(* Logix 5000 project; controller MV vendor 1 type 14 code 217 rev 31.11; software revision 31.00; part 7 of 53 *)
(* tags used below, declared in another part *)
   active : BOOL;
   Ch1_cmd_scan_count : DINT;
   Ch1_DataDelay : TIMER;
   MC_CH1_DRAIN : PlantItem;   // CH1_DRAIN
   MC_CH1_RR : PlantItem;   // CH1_RR
   MC_data_file_value_to_move : DINT;
   MC_N100 : INT[255];   // C1_PLC Channel 1 PLC data
   MC_N101 : INT[255];   // CH1 PC>PLC Channel 1 PC to PLC
   MC_N102 : INT[255];   // CH1 PROG Channel 1 CIP progra m
   MC_N104 : INT[255];   // CH1 REPORT Channel 1 CIP report file
   MC_N108 : INT[255];   // CH1 VDATA Channel 1 CIP progra m validation data
   MC_N120 : INT[255];   // C2 PLC Channel 2 PLC data
   MC_T105 : TIMER[255];   // CH1 TIMERS Channel 1 timers
   MC_T4 : TIMER[255];   // TIMER
(* MC_Common, continued *)

ROUTINE MC_CH1_CMD_101   (* ladder *)
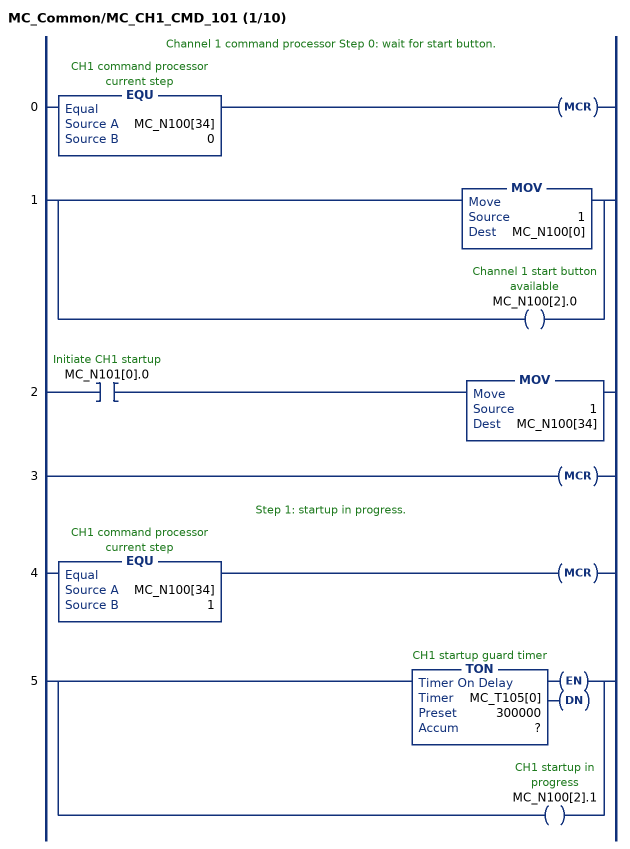
   // Channel 1 command processor Step 0: wait for start button.
   0: EQU(MC_N100[34],0)MCR();
   1: [MOV(1,MC_N100[0]) ,OTE(MC_N100[2].0) ];
   2: XIC(MC_N101[0].0)MOV(1,MC_N100[34]);
   3: MCR();
   // Step 1: startup in progress.
   4: EQU(MC_N100[34],1)MCR();
   5: [TON(MC_T105[0],?,?) ,OTE(MC_N100[2].1) ];
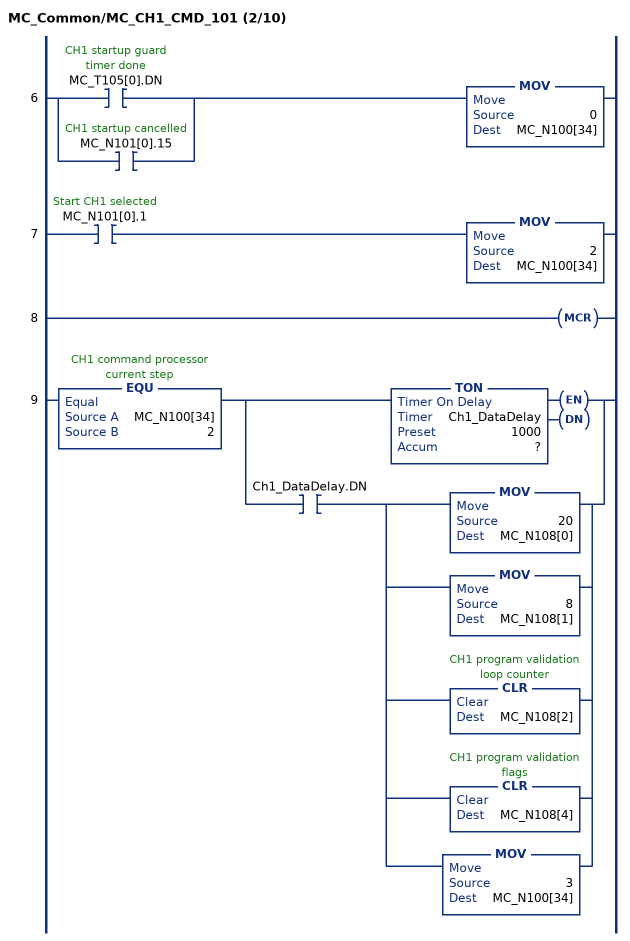
   6: [XIC(MC_T105[0].DN) ,XIC(MC_N101[0].15) ]MOV(0,MC_N100[34]);
   7: XIC(MC_N101[0].1)MOV(2,MC_N100[34]);
   8: MCR();
   9: EQU(MC_N100[34],2)[TON(Ch1_DataDelay,?,?) ,XIC(Ch1_DataDelay.DN) [MOV(20,MC_N108[0]) ,MOV(8,MC_N108[1]) ,CLR(MC_N108[2]) ,CLR(MC_N108[4]) ,MOV(3,MC_N100[34]) ] ];
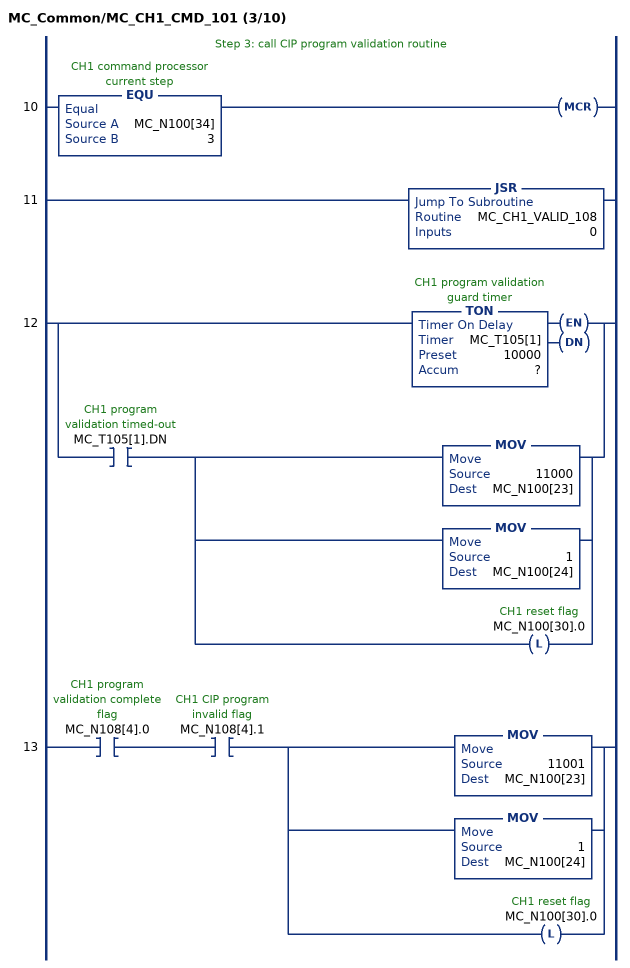
   // Step 3: call CIP program validation routine
   10: EQU(MC_N100[34],3)MCR();
   11: JSR(MC_CH1_VALID_108,0);
   12: [TON(MC_T105[1],?,?) ,XIC(MC_T105[1].DN) [MOV(11000,MC_N100[23]) ,MOV(1,MC_N100[24]) ,OTL(MC_N100[30].0) ] ];
   13: XIC(MC_N108[4].0)XIC(MC_N108[4].1)[MOV(11001,MC_N100[23]) ,MOV(1,MC_N100[24]) ,OTL(MC_N100[30].0) ];
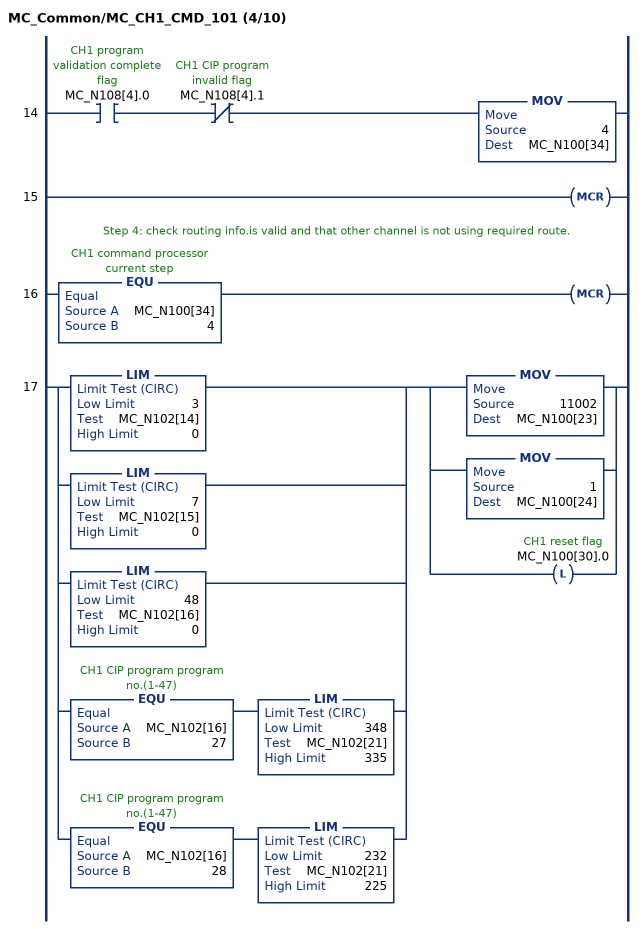
   14: XIC(MC_N108[4].0)XIO(MC_N108[4].1)MOV(4,MC_N100[34]);
   15: MCR();
   // Step 4: check routing info.is valid and that other channel is not using required route.
   16: EQU(MC_N100[34],4)MCR();
   17: [LIM(3,MC_N102[14],0) ,LIM(7,MC_N102[15],0) ,LIM(48,MC_N102[16],0) ,EQU(MC_N102[16],27) LIM(348,MC_N102[21],335) ,EQU(MC_N102[16],28) LIM(232,MC_N102[21],225) ][MOV(11002,MC_N100[23]) ,MOV(1,MC_N100[24]) ,OTL(MC_N100[30].0) ];
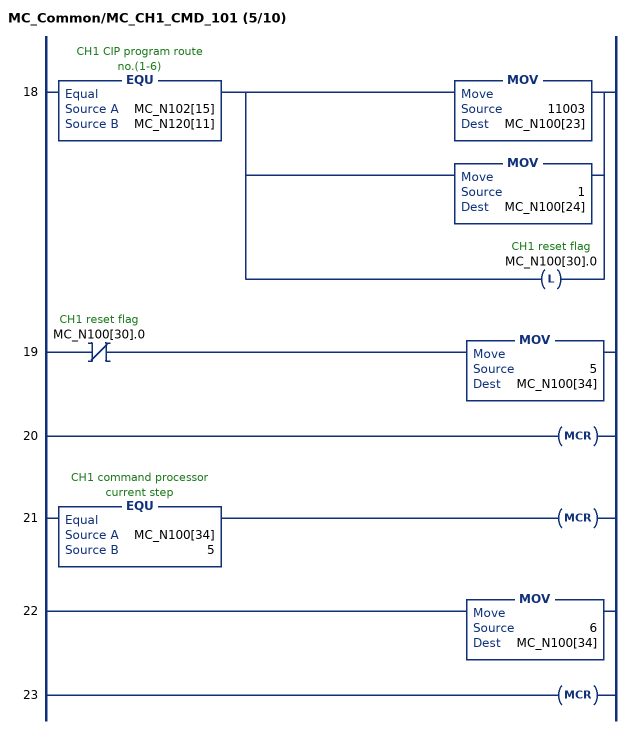
   18: EQU(MC_N102[15],MC_N120[11])[MOV(11003,MC_N100[23]) ,MOV(1,MC_N100[24]) ,OTL(MC_N100[30].0) ];
   19: XIO(MC_N100[30].0)MOV(5,MC_N100[34]);
   20: MCR();
   21: EQU(MC_N100[34],5)MCR();
   22: MOV(6,MC_N100[34]);
   23: MCR();
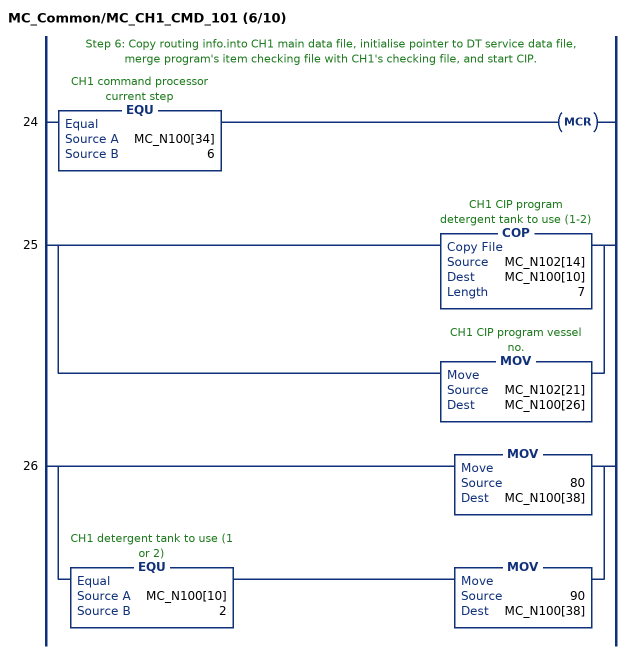
   // Step 6: Copy routing info.into CH1 main data file, initialise pointer to DT service data file, merge program's item checking file with CH1's checking file, and start CIP.
   24: EQU(MC_N100[34],6)MCR();
   25: [COP(MC_N102[14],MC_N100[10],7) ,MOV(MC_N102[21],MC_N100[26]) ];
   26: [MOV(80,MC_N100[38]) ,EQU(MC_N100[10],2) MOV(90,MC_N100[38]) ];
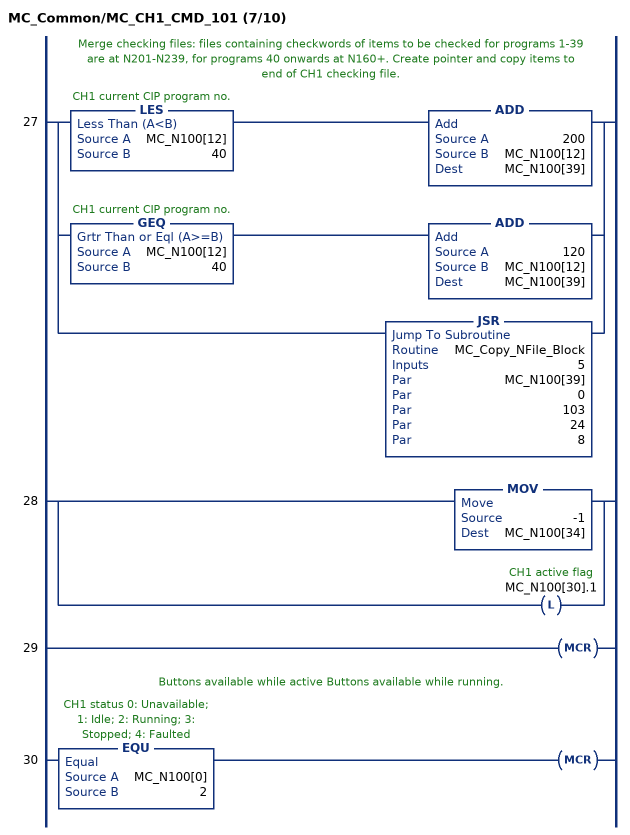
   // Merge checking files: files containing checkwords of items to be checked for programs 1-39 are at N201-N239, for programs 40 onwards at N160+. Create pointer and copy items to end of CH1 checking file.
   27: [LES(MC_N100[12],40) ADD(200,MC_N100[12],MC_N100[39]) ,GEQ(MC_N100[12],40) ADD(120,MC_N100[12],MC_N100[39]) ,JSR(MC_Copy_NFile_Block,5,MC_N100[39],0,103,24,8) ];
   28: [MOV(-1,MC_N100[34]) ,OTL(MC_N100[30].1) ];
   29: MCR();
   // Buttons available while active Buttons available while running.
   30: EQU(MC_N100[0],2)MCR();
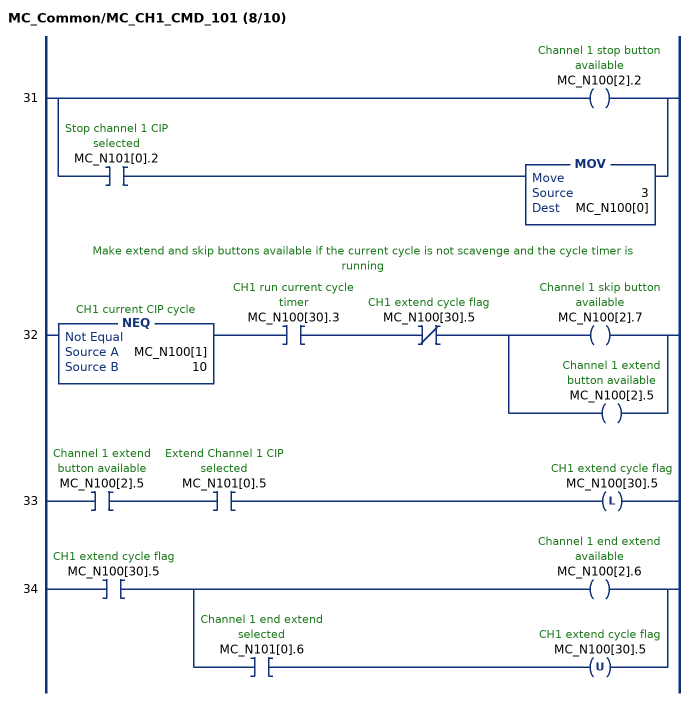
   31: [OTE(MC_N100[2].2) ,XIC(MC_N101[0].2) MOV(3,MC_N100[0]) ];
   // Make extend and skip buttons available if the current cycle is not scavenge and the cycle timer is running
   32: NEQ(MC_N100[1],10)XIC(MC_N100[30].3)XIO(MC_N100[30].5)[OTE(MC_N100[2].7) ,OTE(MC_N100[2].5) ];
   33: XIC(MC_N100[2].5)XIC(MC_N101[0].5)OTL(MC_N100[30].5);
   34: XIC(MC_N100[30].5)[OTE(MC_N100[2].6) ,XIC(MC_N101[0].6) OTU(MC_N100[30].5) ];
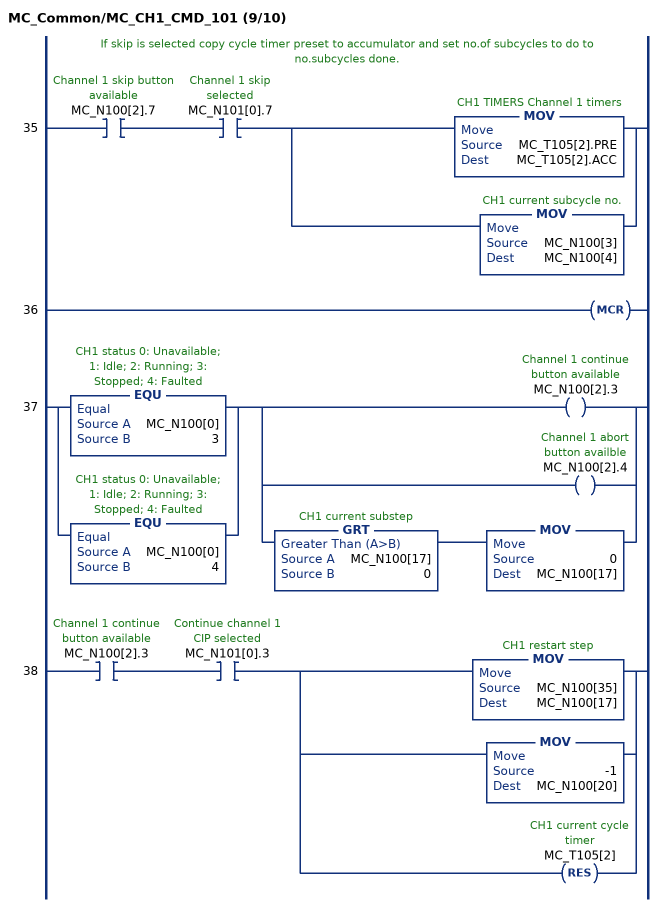
   // If skip is selected copy cycle timer preset to accumulator and set no.of subcycles to do to no.subcycles done.
   35: XIC(MC_N100[2].7)XIC(MC_N101[0].7)[MOV(MC_T105[2].PRE,MC_T105[2].ACC) ,MOV(MC_N100[3],MC_N100[4]) ];
   36: MCR();
   37: [EQU(MC_N100[0],3) ,EQU(MC_N100[0],4) ][OTE(MC_N100[2].3) ,OTE(MC_N100[2].4) ,GRT(MC_N100[17],0) MOV(0,MC_N100[17]) ];
   38: XIC(MC_N100[2].3)XIC(MC_N101[0].3)[MOV(MC_N100[35],MC_N100[17]) ,MOV(-1,MC_N100[20]) ,RES(MC_T105[2]) ];
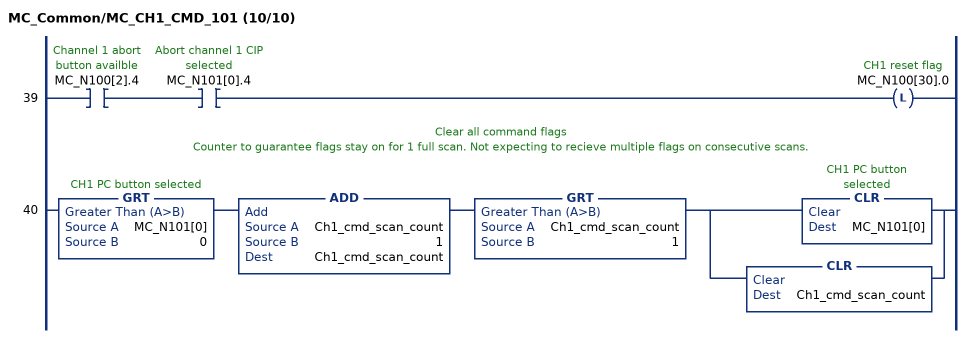
   39: XIC(MC_N100[2].4)XIC(MC_N101[0].4)OTL(MC_N100[30].0);
   // Clear all command flags
   // Counter to guarantee flags stay on for 1 full scan. Not expecting to recieve multiple flags on consecutive scans.
   40: GRT(MC_N101[0],0)ADD(Ch1_cmd_scan_count,1,Ch1_cmd_scan_count)GRT(Ch1_cmd_scan_count,1)[CLR(MC_N101[0]) ,CLR(Ch1_cmd_scan_count) ];
END_ROUTINE

ROUTINE MC_CH1_DETG_112   (* ladder *)
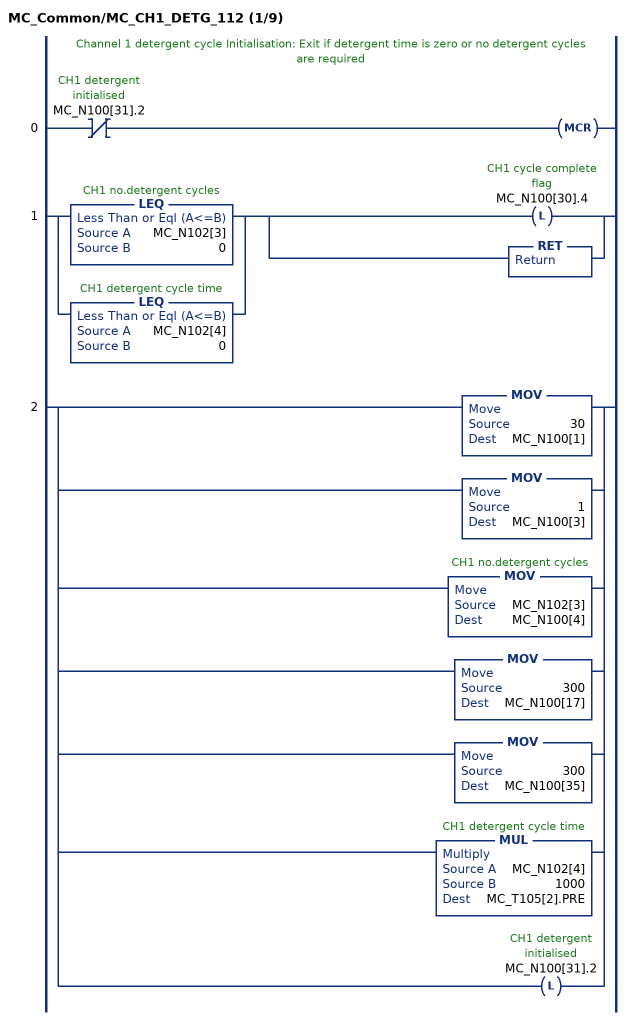
   // Channel 1 detergent cycle Initialisation: Exit if detergent time is zero or no detergent cycles are required
   0: XIO(MC_N100[31].2)MCR();
   1: [LEQ(MC_N102[3],0) ,LEQ(MC_N102[4],0) ][OTL(MC_N100[30].4) ,RET() ];
   2: [MOV(30,MC_N100[1]) ,MOV(1,MC_N100[3]) ,MOV(MC_N102[3],MC_N100[4]) ,MOV(300,MC_N100[17]) ,MOV(300,MC_N100[35]) ,MUL(MC_N102[4],1000,MC_T105[2].PRE) ,OTL(MC_N100[31].2) ];
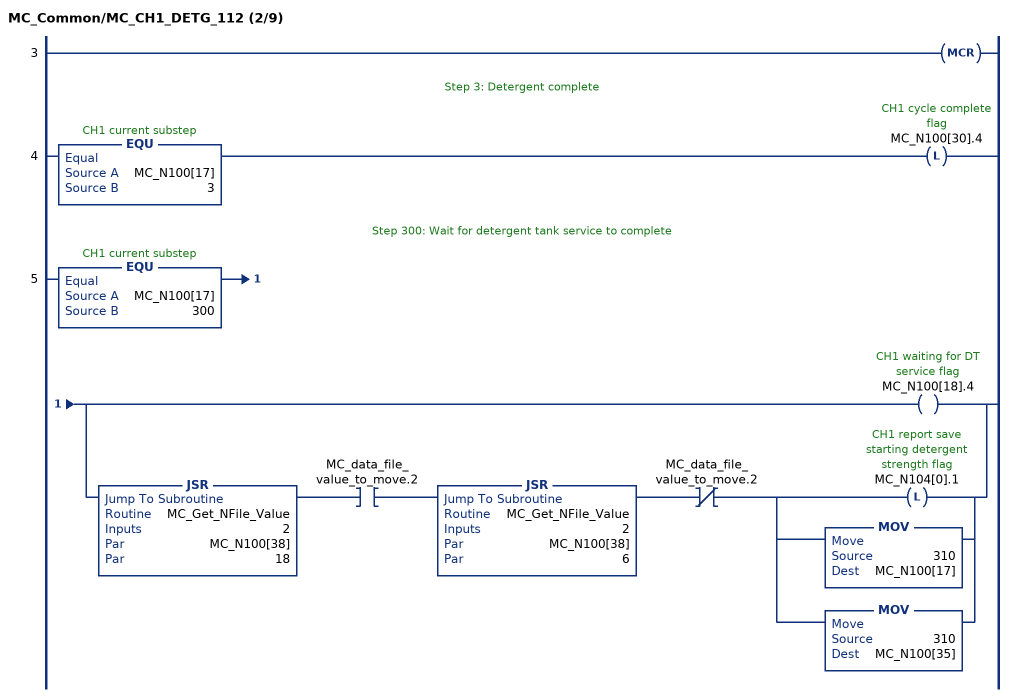
   3: MCR();
   // Step 3: Detergent complete
   4: EQU(MC_N100[17],3)OTL(MC_N100[30].4);
   // Step 300: Wait for detergent tank service to complete
   5: EQU(MC_N100[17],300)[OTE(MC_N100[18].4) ,JSR(MC_Get_NFile_Value,2,MC_N100[38],18) XIC(MC_data_file_value_to_move.2) JSR(MC_Get_NFile_Value,2,MC_N100[38],6) XIO(MC_data_file_value_to_move.2) [OTL(MC_N104[0].1) ,MOV(310,MC_N100[17]) ,MOV(310,MC_N100[35]) ] ];
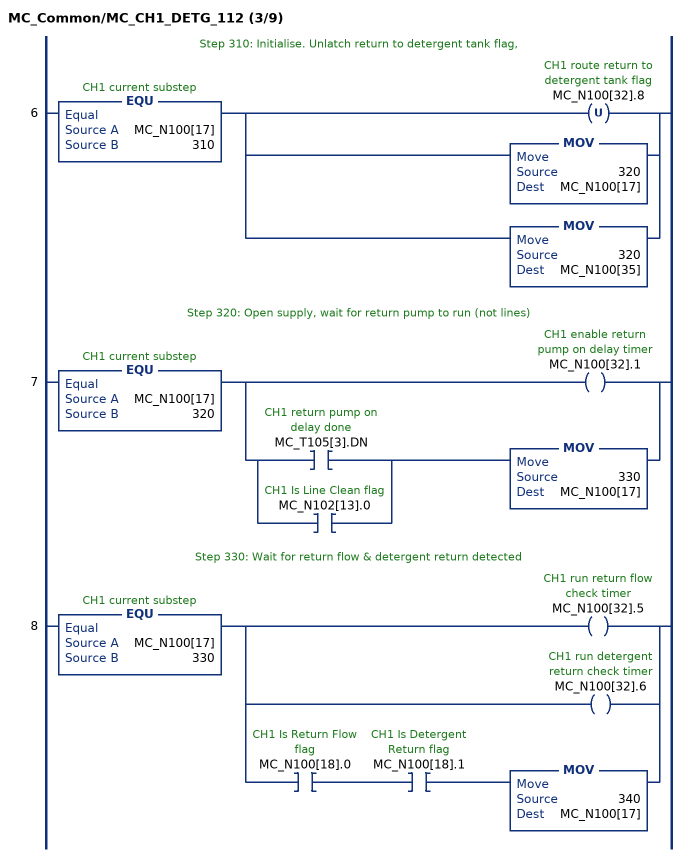
   // Step 310: Initialise. Unlatch return to detergent tank flag,
   6: EQU(MC_N100[17],310)[OTU(MC_N100[32].8) ,MOV(320,MC_N100[17]) ,MOV(320,MC_N100[35]) ];
   // Step 320: Open supply, wait for return pump to run (not lines)
   7: EQU(MC_N100[17],320)[OTE(MC_N100[32].1) ,[XIC(MC_T105[3].DN) ,XIC(MC_N102[13].0) ] MOV(330,MC_N100[17]) ];
   // Step 330: Wait for return flow & detergent return detected
   8: EQU(MC_N100[17],330)[[OTE(MC_N100[32].5) ,OTE(MC_N100[32].6) ] ,XIC(MC_N100[18].0) XIC(MC_N100[18].1) MOV(340,MC_N100[17]) ];
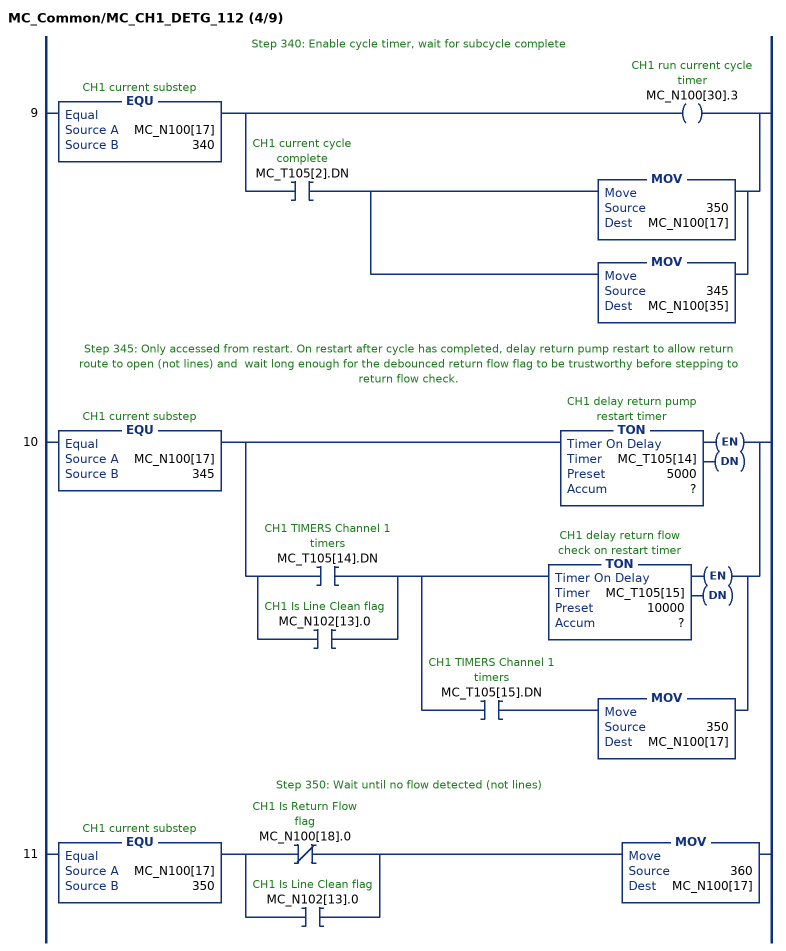
   // Step 340: Enable cycle timer, wait for subcycle complete
   9: EQU(MC_N100[17],340)[OTE(MC_N100[30].3) ,XIC(MC_T105[2].DN) [MOV(350,MC_N100[17]) ,MOV(345,MC_N100[35]) ] ];
   // Step 345: Only accessed from restart. On restart after cycle has completed, delay return pump restart to allow return route to open (not lines) and  wait long enough for the debounced return flow flag to be trustworthy before stepping to return flow check.
   10: EQU(MC_N100[17],345)[TON(MC_T105[14],?,?) ,[XIC(MC_T105[14].DN) ,XIC(MC_N102[13].0) ] [TON(MC_T105[15],?,?) ,XIC(MC_T105[15].DN) MOV(350,MC_N100[17]) ] ];
   // Step 350: Wait until no flow detected (not lines)
   11: EQU(MC_N100[17],350)[XIO(MC_N100[18].0) ,XIC(MC_N102[13].0) ]MOV(360,MC_N100[17]);
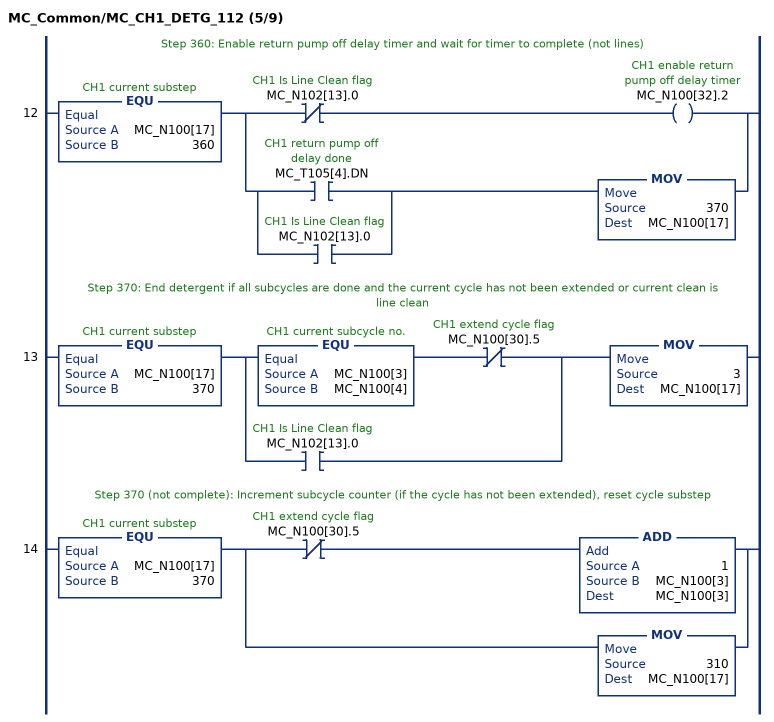
   // Step 360: Enable return pump off delay timer and wait for timer to complete (not lines)
   12: EQU(MC_N100[17],360)[XIO(MC_N102[13].0) OTE(MC_N100[32].2) ,[XIC(MC_T105[4].DN) ,XIC(MC_N102[13].0) ] MOV(370,MC_N100[17]) ];
   // Step 370: End detergent if all subcycles are done and the current cycle has not been extended or current clean is line clean
   13: EQU(MC_N100[17],370)[EQU(MC_N100[3],MC_N100[4]) XIO(MC_N100[30].5) ,XIC(MC_N102[13].0) ]MOV(3,MC_N100[17]);
   // Step 370 (not complete): Increment subcycle counter (if the cycle has not been extended), reset cycle substep
   14: EQU(MC_N100[17],370)[XIO(MC_N100[30].5) ADD(1,MC_N100[3],MC_N100[3]) ,MOV(310,MC_N100[17]) ];
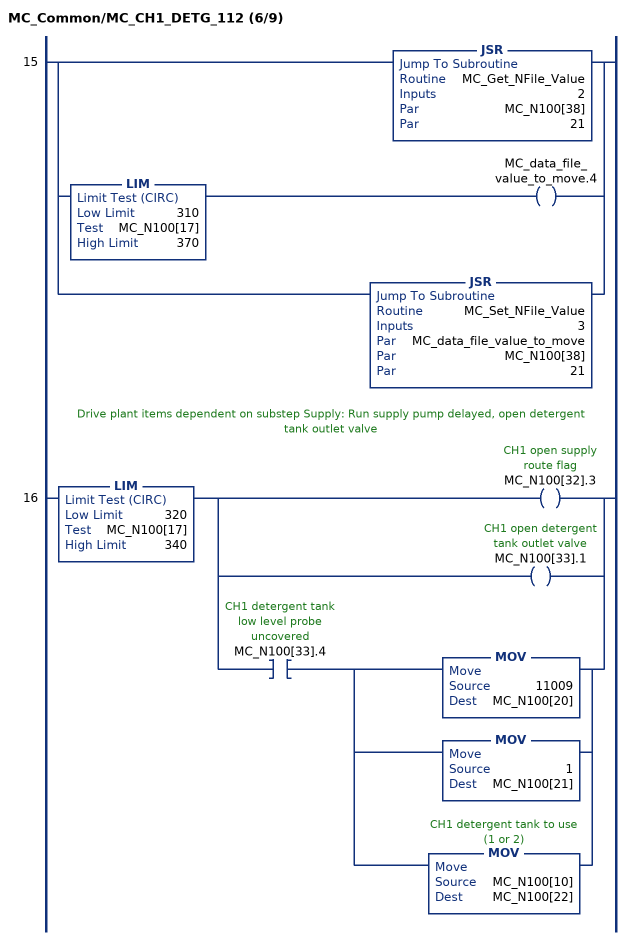
   15: [JSR(MC_Get_NFile_Value,2,MC_N100[38],21) ,LIM(310,MC_N100[17],370) OTE(MC_data_file_value_to_move.4) ,JSR(MC_Set_NFile_Value,3,MC_data_file_value_to_move,MC_N100[38],21) ];
   // Drive plant items dependent on substep Supply: Run supply pump delayed, open detergent tank outlet valve
   16: LIM(320,MC_N100[17],340)[OTE(MC_N100[32].3) ,OTE(MC_N100[33].1) ,XIC(MC_N100[33].4) [MOV(11009,MC_N100[20]) ,MOV(1,MC_N100[21]) ,MOV(MC_N100[10],MC_N100[22]) ] ];
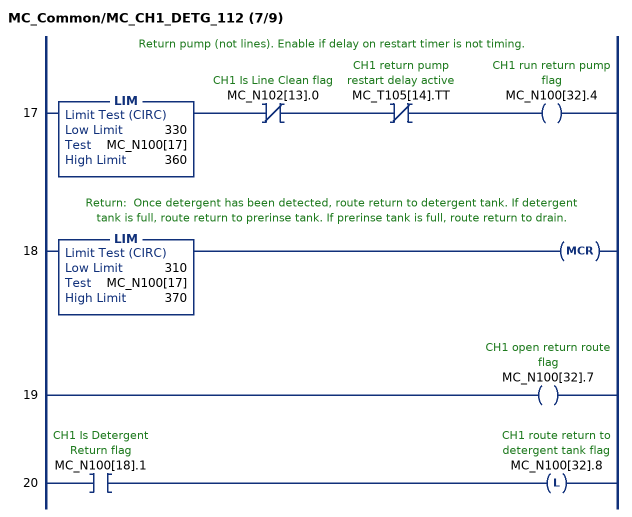
   // Return pump (not lines). Enable if delay on restart timer is not timing.
   17: LIM(330,MC_N100[17],360)XIO(MC_N102[13].0)XIO(MC_T105[14].TT)OTE(MC_N100[32].4);
   // Return:  Once detergent has been detected, route return to detergent tank. If detergent tank is full, route return to prerinse tank. If prerinse tank is full, route return to drain.
   18: LIM(310,MC_N100[17],370)MCR();
   19: OTE(MC_N100[32].7);
   20: XIC(MC_N100[18].1)OTL(MC_N100[32].8);
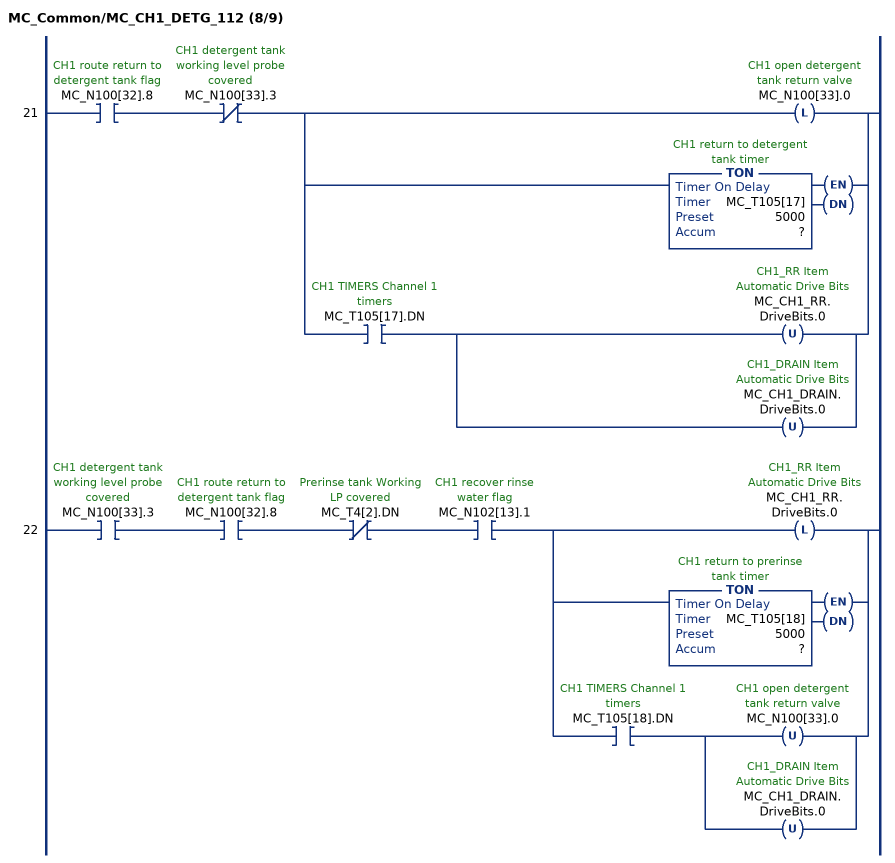
   21: XIC(MC_N100[32].8)XIO(MC_N100[33].3)[OTL(MC_N100[33].0) ,TON(MC_T105[17],?,?) ,XIC(MC_T105[17].DN) [OTU(MC_CH1_RR.DriveBits.0) ,OTU(MC_CH1_DRAIN.DriveBits.0) ] ];
   22: XIC(MC_N100[33].3)XIC(MC_N100[32].8)XIO(MC_T4[2].DN)XIC(MC_N102[13].1)[OTL(MC_CH1_RR.DriveBits.0) ,TON(MC_T105[18],?,?) ,XIC(MC_T105[18].DN) [OTU(MC_N100[33].0) ,OTU(MC_CH1_DRAIN.DriveBits.0) ] ];
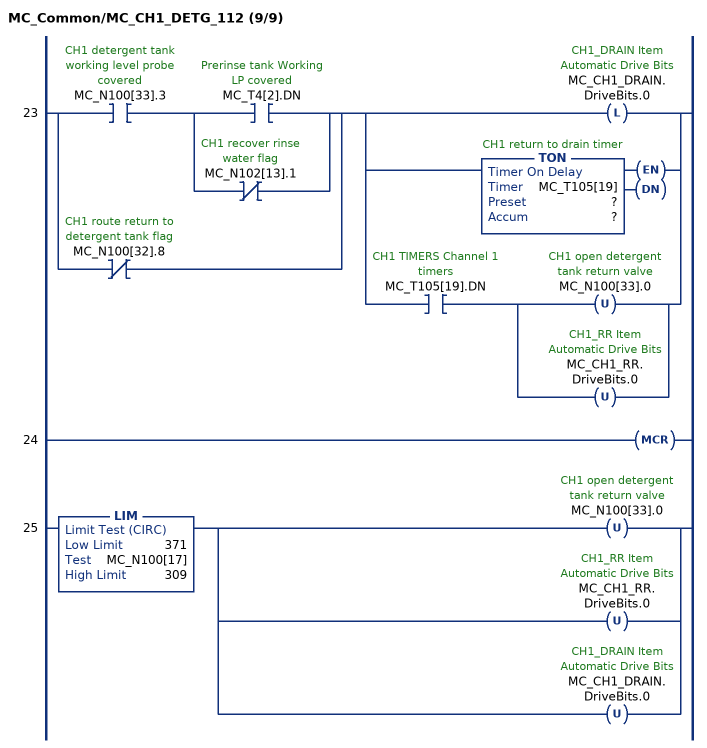
   23: [XIC(MC_N100[33].3) [XIC(MC_T4[2].DN) ,XIO(MC_N102[13].1) ] ,XIO(MC_N100[32].8) ][OTL(MC_CH1_DRAIN.DriveBits.0) ,TON(MC_T105[19],?,?) ,XIC(MC_T105[19].DN) [OTU(MC_N100[33].0) ,OTU(MC_CH1_RR.DriveBits.0) ] ];
   24: MCR();
   25: LIM(371,MC_N100[17],309)[OTU(MC_N100[33].0) ,OTU(MC_CH1_RR.DriveBits.0) ,OTU(MC_CH1_DRAIN.DriveBits.0) ];
END_ROUTINE
